// TIA Portal project "oscat_basic_332_s7_TIA_V12_V13_SP1_V14_V15.1" (V15.1)

(* hardware
DEVICE "Rack 0"  S7-300 station
   slot 0: "Profilschiene_0"  Rail  6ES7 390-1***0-0AA0
   slot 2: "Buffer Management"  Unspecific CPU S7 300  6ES7 3XX-XXXXX-XXXX
DEVICE "Rack 0_2"  S7-300 station
   slot 0: "Profilschiene_0"  Rail  6ES7 390-1***0-0AA0
   slot 2: "Constants"  Unspecific CPU S7 300  6ES7 3XX-XXXXX-XXXX
DEVICE "Rack 0_3"  S7-300 station
   slot 0: "Profilschiene_0"  Rail  6ES7 390-1***0-0AA0
   slot 2: "Eng signal generators"  Unspecific CPU S7 300  6ES7 3XX-XXXXX-XXXX
DEVICE "Rack 0_4"  S7-300 station
   slot 0: "Profilschiene_0"  Rail  6ES7 390-1***0-0AA0
   slot 2: "Eng signal processing"  Unspecific CPU S7 300  6ES7 3XX-XXXXX-XXXX
DEVICE "Rack 0_5"  S7-300 station
   slot 0: "Profilschiene_0"  Rail  6ES7 390-1***0-0AA0
   slot 2: "Engineering automation"  Unspecific CPU S7 300  6ES7 3XX-XXXXX-XXXX
DEVICE "Rack 0_6"  S7-300 station
   slot 0: "Profilschiene_0"  Rail  6ES7 390-1***0-0AA0
   slot 2: "Engineering control"  Unspecific CPU S7 300  6ES7 3XX-XXXXX-XXXX
DEVICE "Rack 0_7"  S7-300 station
   slot 0: "Profilschiene_0"  Rail  6ES7 390-1***0-0AA0
   slot 2: "Engineering conversion"  Unspecific CPU S7 300  6ES7 3XX-XXXXX-XXXX
DEVICE "Rack 0_8"  S7-300 station
   slot 0: "Profilschiene_0"  Rail  6ES7 390-1***0-0AA0
   slot 2: "Engineering measurements"  Unspecific CPU S7 300  6ES7 3XX-XXXXX-XXXX
DEVICE "Rack 0_9"  S7-300 station
   slot 0: "Profilschiene_0"  Rail  6ES7 390-1***0-0AA0
   slot 2: "Engineering sensor"  Unspecific CPU S7 300  6ES7 3XX-XXXXX-XXXX
DEVICE "Rack 0_10"  S7-300 station
   slot 0: "Profilschiene_0"  Rail  6ES7 390-1***0-0AA0
   slot 2: "List Processing"  Unspecific CPU S7 300  6ES7 3XX-XXXXX-XXXX
DEVICE "Rack 0_11"  S7-300 station
   slot 0: "Profilschiene_0"  Rail  6ES7 390-1***0-0AA0
   slot 2: "Logic FF edge triggered"  Unspecific CPU S7 300  6ES7 3XX-XXXXX-XXXX
DEVICE "Rack 0_12"  S7-300 station
   slot 0: "Profilschiene_0"  Rail  6ES7 390-1***0-0AA0
   slot 2: "Logic FF pulse triggered"  Unspecific CPU S7 300  6ES7 3XX-XXXXX-XXXX
DEVICE "Rack 0_13"  S7-300 station
   slot 0: "Profilschiene_0"  Rail  6ES7 390-1***0-0AA0
   slot 2: "Logic Others"  Unspecific CPU S7 300  6ES7 3XX-XXXXX-XXXX
DEVICE "Rack 0_14"  S7-300 station
   slot 0: "Profilschiene_0"  Rail  6ES7 390-1***0-0AA0
   slot 2: "Logic gate logic"  Unspecific CPU S7 300  6ES7 3XX-XXXXX-XXXX
DEVICE "Rack 0_15"  S7-300 station
   slot 0: "Profilschiene_0"  Rail  6ES7 390-1***0-0AA0
   slot 2: "Logic generators"  Unspecific CPU S7 300  6ES7 3XX-XXXXX-XXXX
DEVICE "Rack 0_16"  S7-300 station
   slot 0: "Profilschiene_0"  Rail  6ES7 390-1***0-0AA0
   slot 2: "Logic memory"  Unspecific CPU S7 300  6ES7 3XX-XXXXX-XXXX
DEVICE "Rack 0_17"  S7-300 station
   slot 0: "Profilschiene_0"  Rail  6ES7 390-1***0-0AA0
   slot 2: "Math Double Precision"  Unspecific CPU S7 300  6ES7 3XX-XXXXX-XXXX
DEVICE "Rack 0_18"  S7-300 station
   slot 0: "Profilschiene_0"  Rail  6ES7 390-1***0-0AA0
   slot 2: "Math Vektormathematik"  Unspecific CPU S7 300  6ES7 3XX-XXXXX-XXXX
DEVICE "Rack 0_19"  S7-300 station
   slot 0: "Profilschiene_0"  Rail  6ES7 390-1***0-0AA0
   slot 2: "Mathematical"  Unspecific CPU S7 300  6ES7 3XX-XXXXX-XXXX
DEVICE "Rack 0_20"  S7-300 station
   slot 0: "Profilschiene_0"  Rail  6ES7 390-1***0-0AA0
   slot 2: "Mathematical Array"  Unspecific CPU S7 300  6ES7 3XX-XXXXX-XXXX
DEVICE "Rack 0_21"  S7-300 station
   slot 0: "Profilschiene_0"  Rail  6ES7 390-1***0-0AA0
   slot 2: "Mathematical Complex"  Unspecific CPU S7 300  6ES7 3XX-XXXXX-XXXX
DEVICE "Rack 0_22"  S7-300 station
   slot 0: "Profilschiene_0"  Rail  6ES7 390-1***0-0AA0
   slot 2: "Mathematical Geometry"  Unspecific CPU S7 300  6ES7 3XX-XXXXX-XXXX
DEVICE "Rack 0_23"  S7-300 station
   slot 0: "Profilschiene_0"  Rail  6ES7 390-1***0-0AA0
   slot 2: "Mathematical functions"  Unspecific CPU S7 300  6ES7 3XX-XXXXX-XXXX
DEVICE "Rack 0_24"  S7-300 station
   slot 0: "Profilschiene_0"  Rail  6ES7 390-1***0-0AA0
   slot 2: "Other"  Unspecific CPU S7 300  6ES7 3XX-XXXXX-XXXX
DEVICE "Rack 0_25"  S7-300 station
   slot 0: "Profilschiene_0"  Rail  6ES7 390-1***0-0AA0
   slot 2: "String"  Unspecific CPU S7 300  6ES7 3XX-XXXXX-XXXX
DEVICE "Rack 0_26"  S7-300 station
   slot 0: "Profilschiene_0"  Rail  6ES7 390-1***0-0AA0
   slot 2: "Time and Date"  Unspecific CPU S7 300  6ES7 3XX-XXXXX-XXXX
DEVICE "Rack 0_27"  S7-300 station
   slot 0: "Profilschiene_0"  Rail  6ES7 390-1***0-0AA0
   slot 2: "xS7"  Unspecific CPU S7 300  6ES7 3XX-XXXXX-XXXX
*)

// ===== PLC "Buffer Management"  Unspecific CPU S7 300 =====

DATA_BLOCK "SETUP"   // DB1
TITLE = SETUP
{ S7_Optimized_Access := 'FALSE' }
AUTHOR : oscat
FAMILY : CONSTANT
NAME : DBSETUP
VERSION : 1.0
   VAR
      EXTENDED_ASCII : Bool := TRUE;
      CHARNAMES : Array[1..4] of String[253];
      MTH_OFS : Array[1..12] of Int;
      DECADES : Array[0..8] of Real;
   END_VAR
BEGIN
   CHARNAMES[1] := ';"&quot;&&amp;<&lt;>&gt;€&euro; &nbsp;¡&iexcl;¢&cent;£&pound;¤&curren;¥&yen;¦&brvbar;§&sect;¨&uml;©&copy;ª&ordf;«&laquo;¬&not;­&shy;®&reg;¯&macr;°&deg;±&plusmn;²&sup2;³&sup3;´&acute;µ&micro;¶&para;·&middot;¸&cedil;¹&sup1;º&ordm;»&raquo;¼&frac14;Û&Ucirc;';
   CHARNAMES[2] := ';¾&frac34;¿&iquest;À&Agrave;Á&Aacute;Â&Acirc;Ã&Atilde;Ä&Auml;Å&Aring;Æ&AElig;Ç&Ccedil;È&Egrave;É&Eacute;Ê&Ecirc;Ë&Euml;Ì&Igrave;Í&Iacute;Î&Icirc;Ï&Iuml;Ð&ETH;Ñ&Ntilde;Ò&Ograve;Ó&Oacute;Ô&Ocirc;Õ&Otilde;Ö&Ouml;×&times;Ø&Oslash;Ù&Ugrave;Ú&Uacute;½&frac12;';
   CHARNAMES[3] := ';Ü&Uuml;Ý&Yacute;Þ&THORN;ß&szlig;à&agrave;á&aacute;â&acirc;ã&atilde;ä&auml;å&aring;æ&aelig;ç&ccedil;è&egrave;é&eacute;ê&ecirc;ë&euml;ì&igrave;í&iacute;î&icirc;ï&iuml;ð&eth;ñ&ntilde;ò&ograve;ó&oacute;ô&ocirc;õ&otilde;ö&ouml;÷&divide;ø&oslash;ù&ugrave;';
   CHARNAMES[4] := ';ú&uacute;û&ucirc;ü&uuml;ý&yacute;þ&thorn;ÿ&yuml;';
   MTH_OFS[2] := 31;
   MTH_OFS[3] := 59;
   MTH_OFS[4] := 90;
   MTH_OFS[5] := 120;
   MTH_OFS[6] := 151;
   MTH_OFS[7] := 181;
   MTH_OFS[8] := 212;
   MTH_OFS[9] := 243;
   MTH_OFS[10] := 273;
   MTH_OFS[11] := 304;
   MTH_OFS[12] := 334;
   DECADES[0] := 1.0e+0;
   DECADES[1] := 1.0e+1;
   DECADES[2] := 1.0e+2;
   DECADES[3] := 1.0e+3;
   DECADES[4] := 1.0e+4;
   DECADES[5] := 1.0e+4;
   DECADES[6] := 1.0e+5;
   DECADES[7] := 1.0e+6;
   DECADES[8] := 1.0e+7;
END_DATA_BLOCK

FUNCTION_BLOCK "_BUFFER_CLEAR"   // FB225, SCL
TITLE = _BUFFER_CLEAR
{ S7_Optimized_Access := 'FALSE' }
AUTHOR : hugo
FAMILY : BUFFER
NAME : BCLEAR
VERSION : 1.2
// this function will initialize a given array of byte with 0.
// the function needs to be called:    _buffer_clear(adr("array"),sizeof("array"));
// this function will manipulate a given array.
// the function manipulates the original array, it rerturnes true when finished.
// because this function works with pointers its very time efficient and it needs no extra memory.
   VAR_INPUT
      PT : Pointer;
      _PT AT PT : Struct
         DBNr : Word;
         Adr : DWord;
      END_STRUCT;
      SIZE : Int;
   END_VAR
   VAR_OUTPUT
      _CLEAR : Bool;
   END_VAR
   VAR_TEMP
      ptw : Int;   // POINTER TO DWORD;
      temp : DWord;
      end : DWord;
      end32 : DWord;
      tPT : Int;
   END_VAR
BEGIN


   #_CLEAR := FALSE;

   #tPT := DWORD_TO_INT(SHR(IN:=SHL(IN:=#_PT.Adr,N:=8),N:=11));

   (* this routine uses 32 bit access to gain speed *)
   (* first access bytes till pointer is aligned for 32 bit access *)
   #temp := INT_TO_DWORD(#tPT);  //pt;
   #end := DINT_TO_DWORD(DWORD_TO_DINT(#temp) + #SIZE);
   #end32 := DINT_TO_DWORD(DWORD_TO_DINT(#end) - 4);   //end32 := end - 3;
   WHILE (#tPT < DWORD_TO_DINT(#end)) AND (DWORD_TO_DINT((#temp AND 16#00000003)) > 0) DO
       WORD_TO_BLOCK_DB(#_PT.DBNr).DB(#tPT) := 0;
       #tPT := #tPT + 1;
       #temp := DINT_TO_DWORD(DWORD_TO_DINT(#temp) + 1);
   END_WHILE;
   (* pointer is aligned, now copy 32 bits at a time *)
   #ptw := #tPT;
   WHILE #ptw < DWORD_TO_DINT(#end32) DO
       WORD_TO_BLOCK_DB(#_PT.DBNr).DD(#ptw) := 0;
       #ptw := #ptw + 4;
   END_WHILE;
   (* copy the remaining bytes in byte mode *)
   #tPT := #ptw;    //ptw;
   WHILE #tPT < DWORD_TO_DINT(#end) DO
       WORD_TO_BLOCK_DB(#_PT.DBNr).DB(#tPT) := 0;
       #tPT := #tPT + 1;
   END_WHILE;

   #_CLEAR := TRUE;

   (* revision History
   hm  5. mar. 2008    rev 1.0
       original version

   hm  16. mar. 2008   rev 1.1
       added type conversion to avoid warnings under codesys 30
       chaged type of input size to uint
       deleted unused variable i

   hm  31. oct. 2008   rev 1.2
       corrected an error while routine would write outside of arrays

   *)
END_FUNCTION_BLOCK

FUNCTION_BLOCK "_BUFFER_INIT"   // FB226, SCL
TITLE = _BUFFER_INIT
{ S7_Optimized_Access := 'FALSE' }
AUTHOR : hugo
FAMILY : BUFFER
NAME : BINIT
VERSION : 1.2
// this function will initialize a given array of byte with init.
// the function needs to be called:    _buffer_init(adr("array"),sizeof("array"),init);
// this function will manipulate a given array.
// the function manipulates the original array, it rerturnes true when finished.
// because this function works with pointers its very time efficient and it needs no extra memory.
   VAR_INPUT
      pt : Pointer;
      _pt AT pt : Struct
         DBNr : Word;
         Adr : DWord;
      END_STRUCT;
      size : Int;
      init : Byte;
   END_VAR
   VAR_OUTPUT
      _INIT : Bool;
   END_VAR
   VAR_TEMP
      ptw : Int;   // ptw : POINTER TO DWORD;
      temp : DWord;
      end : DWord;
      end32 : DWord;
      tPT : Int;
   END_VAR
BEGIN


   #_INIT := FALSE;
   #tPT := DWORD_TO_INT(SHR(IN:=SHL(IN:=#_pt.Adr,N:=8),N:=11));

   (* this routine uses 32 bit access to gain speed *)
   (* first access bytes till pointer is aligned for 32 bit access *)
   #temp := INT_TO_DWORD(#tPT);
   #end := DINT_TO_DWORD(DWORD_TO_DINT(#temp) + #size);
   #end32 := DINT_TO_DWORD(DWORD_TO_DINT(#temp) - 4);    //end32 := end - 3;
   WHILE (#tPT < DWORD_TO_DINT(#end)) AND (DWORD_TO_DINT((#temp AND 16#00000003)) > 0) DO
       WORD_TO_BLOCK_DB(#_pt.DBNr).DB(#tPT) := #init;
       #tPT := #tPT + 1;
       #temp := DINT_TO_DWORD(DWORD_TO_DINT(#temp) + 1);
   END_WHILE;
   (* pointer is aligned, now copy 32 bits at a time *)
   #ptw := #tPT;
   #temp := SHL(IN:=BYTE_TO_DWORD(#init),N:=24) OR SHL(IN:=BYTE_TO_DWORD(#init),N:=16) OR SHL(IN:=BYTE_TO_DWORD(#init),N:=8) OR BYTE_TO_DWORD(#init);
   WHILE #ptw < DWORD_TO_DINT(#end32) DO
       WORD_TO_BLOCK_DB(#_pt.DBNr).DD(#ptw) := #temp;
       #ptw := #ptw + 4;
   END_WHILE;
   (* copy the remaining bytes in byte mode *)
   #tPT := #ptw;
   WHILE #tPT < DWORD_TO_DINT(#end) DO
       WORD_TO_BLOCK_DB(#_pt.DBNr).DB(#tPT) := #init;
       #tPT := #tPT + 1;
   END_WHILE;

   #_INIT := TRUE;

   (* revision History
   hm  5. mar. 2008    rev 1.0
       original version

   hm  16. mar. 2008   rev 1.1
       added type conversion to avoid warnings under codesys 3.0
       chaged type of input size to uint.

   hm  31. oct. 2008   rev 1.2
       corrected an error while routine would write outside of arrays

   *)
END_FUNCTION_BLOCK

FUNCTION_BLOCK "_BUFFER_INSERT"   // FB227, SCL
TITLE = _BUFFER_INSERT
{ S7_Optimized_Access := 'FALSE' }
AUTHOR : hugo
FAMILY : BUFFER
NAME : BINSERT
VERSION : 1.4
// this function will initialize a given array of byte with init.
// the function needs to be called:    _buffer_init(adr("array"),sizeof("array"),init);
// this function will manipulate a given array.
// the function manipulates the original array, it rerturnes true when finished.
// because this function works with pointers its very time efficient and it needs no extra memory.
// 
// uses: STRING_TO_BUFFER [FB228]
   VAR_INPUT
      STR : String[254];
      _str AT STR : Struct
         length : Byte;
         act_length : Byte;
         str : Array[1..254] of Byte;
      END_STRUCT;
      POS : Int;
      PT : Pointer;
      _pt AT PT : Struct
         DBNr : Word;
         Adr : DWord;
      END_STRUCT;
      SIZE : Int;
   END_VAR
   VAR_OUTPUT
      OUT : Bool;
   END_VAR
   VAR
      STRING_TO_BUFFER : "_STRING_TO_BUFFER";
   END_VAR
   VAR_TEMP
      end : Int;
      lx : Int;
      i : Int;
      tPT : Int;
   END_VAR
BEGIN


   #OUT := FALSE;

   #tPT := DWORD_TO_INT(SHR(IN:=SHL(IN:=#_pt.Adr,N:=8),N:=11));

   #POS := LIMIT(MN:=0,IN:=#POS,MX:=#SIZE - 1);
   #lx := BYTE_TO_INT(#_str.length);  //LEN(str);
   #end := #POS + #lx;
   (* first move the upper part of the buffer to make space for the string *)
   FOR #i := #SIZE - 1 TO #end BY -1 DO
       WORD_TO_BLOCK_DB(#_pt.DBNr).DB(#tPT+#i) := WORD_TO_BLOCK_DB(#_pt.DBNr).DB(#tPT+#i-#lx);
   END_FOR;
   (* copy the string *)
   #STRING_TO_BUFFER(strBLKMOV#STR, pos:=#POS, pt:=#PT, size:=#SIZE);
   #OUT := #STRING_TO_BUFFER._BUFFER;


   (* revision History
   hm  9. mar. 2008  rev 1.0
     original version

   hm  16. mar. 2008 rev 1.1
     changed type of input size to uint

   hm  13. may. 2008 rev 1.2
     changed type of pointer to array[1..32767]
     changed size of string to STRING_LENGTH

   hm  23. mar. 2009 rev 1.3
     avoid writing to input pos

   hm  12. nov. 2009 rev 1.4
     code optimized

   *)
END_FUNCTION_BLOCK

FUNCTION_BLOCK "_STRING_TO_BUFFER"   // FB228, SCL
TITLE = _STRING_TO_BUFFER
{ S7_Optimized_Access := 'FALSE' }
AUTHOR : hugo
FAMILY : BUFFER
NAME : BSTRB
VERSION : 1.3
// this function will copy a string into an array of byte starting at position pos.
// the function needs to be called:    _String_To_buffer(str, pos, adr("array"),sizeof("array"));
// this function will manipulate the array directly in memory and returns true when finished.
// because this function works with pointers its very time efficient and it needs no extra memory.
   VAR_INPUT
      str : String[254];
      _str AT str : Struct
         length : Byte;
         act_length : Byte;
         str : Array[1..254] of Byte;
      END_STRUCT;
      pos : Int;
      pt : Pointer;
      _pt AT pt : Struct
         DBNr : Word;
         Adr : DWord;
      END_STRUCT;
      size : Int;
   END_VAR
   VAR_OUTPUT
      _BUFFER : Bool;
   END_VAR
   VAR_TEMP
      ps : Int;   // POINTER TO BYTE;
      i : Int;
      end : Int;
      tPT : Int;
   END_VAR
BEGIN


   #_BUFFER := FALSE;
   #tPT := DWORD_TO_INT(SHR(IN:=SHL(IN:=#_pt.Adr,N:=8),N:=11));

   #ps := 1;    //ADR(str);
   #end := MIN(IN1:=#pos + BYTE_TO_INT(#_str.length) - 1,IN2:=#size);
   IF #end > 0 THEN #end := #end -1; END_IF;
   FOR #i := #pos TO #end DO
       WORD_TO_BLOCK_DB(#_pt.DBNr).DB(#tPT+#i-1) := #_str.str[#ps];
       #ps := #ps + 1;
   END_FOR;

   #_BUFFER := TRUE;

   (* revision History

   hm  5. mar. 2008 rev 1.0
    original version

   hm 16. mar. 2008 rev 1.1
    changed type of input size to uint

   hm 13. may. 2008 rev 1.2
    changed type of pointer to array[1..32767]
    changed size of string to STRING_LENGTH

   hm 12. nov. 2009 rev 1.3
    limit end to size - 1

   *)
END_FUNCTION_BLOCK

FUNCTION_BLOCK "BUFFER_SEARCH"   // FB229, SCL
TITLE = BUFFER_SEARCH
{ S7_Optimized_Access := 'FALSE' }
AUTHOR : hugo
FAMILY : BUFFER
NAME : BSEARCH
VERSION : 1.4
// this function will search for a string STR in an array of byte starting at position pos.
// the function needs to be called: buffer_search(adr("array"),sizeof("array"), STR, POS, IGN);
// because this function works with pointers its very time efficient and it needs no extra memory.
// The function returns the position of the first character of the string in the array if found.
// a -1 is returned if the string is not found in the array.
// when IGN = TRUE, STR must be in capital letters and the search is case insensitv.
   VAR_INPUT
      PT : Pointer;
      _pt AT PT : Struct
         DBNr : Word;
         Adr : DWord;
      END_STRUCT;
      SIZE : Int;
      STR : String[254];
      _str AT STR : Struct
         length : Byte;
         act_length : Byte;
         str : Array[1..254] of Byte;
      END_STRUCT;
      POS : Int;
      IGN : Bool;
   END_VAR
   VAR_OUTPUT
      _SEARCH : Int;
   END_VAR
   VAR_TEMP
      ps : Int;   // POINTER TO ARRAY[0..255] OF BYTE;
      chx : Byte;
      i : Int;
      end : Int;
      k : Int;
      lx : Int;
      tPT : Int;
   END_VAR
BEGIN


   #tPT := DWORD_TO_INT(SHR(IN:=SHL(IN:=#_pt.Adr,N:=8),N:=11));

   #ps := 1;    //ADR(str);
   #lx := BYTE_TO_INT(#_str.act_length);  //LEN(str);
   #end := MIN(IN1:=#SIZE - #lx, IN2:= #SIZE - 1);
   #lx := #lx - 1;
   FOR #i := #POS TO #end DO
     FOR #k := 0 TO #lx DO
       //IF (_str.str[ps+k] <> ign) AND (_str.str[ps+k] <> WORD_TO_BLOCK_DB(_pt.DBNr).DB[tPT+i+k]) THEN EXIT; END_IF;
       IF #IGN THEN 
         #chx := "TO_UPPER"(WORD_TO_BLOCK_DB(#_pt.DBNr).DB(#tPT+#i+#k)); 
       ELSE 
         #chx := WORD_TO_BLOCK_DB(#_pt.DBNr).DB(#tPT+#i+#k); 
       END_IF;
       IF WORD_TO_BLOCK_DB(#_pt.DBNr).DB(#tPT+#k) <> #chx THEN 
         EXIT; 
       END_IF;
     END_FOR;
     IF #k > #lx THEN
       #_SEARCH := #i;
       RETURN;
     END_IF;
   END_FOR;
   #_SEARCH := -1;


   (* revision History

   hm 5. mar. 2008 rev 1.0
     original version

   hm  16. mar. 2008 rev 1.1
     chaged type of input size to uint

   hm  13. may. 2008 rev 1.2
     changed type of pointer to array[1..32767]
     changed size of string to STRING_LENGTH

   hm  12. nov. 2009 rev 1.3
     limit end to array size

   hm  25. jan. 2011 rev 1.4
     ign = True will now ignore case
     return -1 if nothing found
   *)
END_FUNCTION_BLOCK

FUNCTION_BLOCK "BUFFER_TO_STRING"   // FB230, SCL
TITLE = BUFFER_TO_STRING
{ S7_Optimized_Access := 'FALSE' }
AUTHOR : hugo
FAMILY : BUFFER
NAME : BBSTR
VERSION : 1.5
// this function will retrieve a string from an array of byte starting at position start and stop at position stop.
// the function needs to be called: buffer_TO_String(adr("array"),sizeof("array"), start, stop);
// because this function works with pointers its very time efficient and it needs no extra memory.
   VAR_INPUT
      PT : Pointer;
      _pt AT PT : Struct
         DBNr : Word;
         Adr : DWord;
      END_STRUCT;
      SIZE : Int;
      START : Int;
      STOP : Int;
   END_VAR
   VAR_OUTPUT
      _STRING : String[254];
      _str AT _STRING : Struct
         length : Byte;
         act_length : Byte;
         str : Array[1..254] of Byte;
      END_STRUCT;
   END_VAR
   VAR_TEMP
      ps : Int;   // POINTER TO BYTE;
      i : Int;
      tPT : Int;
      stp : Int;
      sta : Int;
   END_VAR
BEGIN


   #tPT := DWORD_TO_INT(SHR(IN:=SHL(IN:=#_pt.Adr,N:=8),N:=11));

   #ps := 1;    //ADR(BUFFER_TO_STRING);
   IF #SIZE = 0 THEN RETURN; END_IF;
   #sta := MIN(IN1:=#START, IN2:=#SIZE-1);
   #stp := MIN(IN1:=#STOP, IN2:=#SIZE-1);

   (* check for maximum string_length *)
   IF (#stp - #sta + 1) >= BYTE_TO_INT(#_str.act_length) THEN
     #stp := #sta + BYTE_TO_INT(#_str.act_length) - 1;
   END_IF;

   FOR #i := #sta TO #stp DO
       #_str.str[#ps] := WORD_TO_BLOCK_DB(#_pt.DBNr).DB(#tPT+#i);
       #ps := #ps + 1;
   END_FOR;

   (* terminate the string *)
   #_str.act_length := INT_TO_BYTE(#ps-1);

   (* revision History
   hm  5. mar. 2008  rev 1.0
     original version

   hm  16. mar. 2008 rev 1.1
     changed type of input size to uint

   hm  13. may. 2008 rev 1.2
     changed type of pointer to array[0..32767]
     changed size of string to STRING_LENGTH

   hm  12. jun. 2008 rev 1.3
     check for pointer overrun
     change input start and stop to uint
     added type conversions to avoid warnings under codesys 3.0

   hm  23. mar. 2009 rev 1.4
     avoid writing to input stop

   hm  12. nov. 2009 rev 1.5
     limit start and stop to size -1

   *)
END_FUNCTION_BLOCK

FUNCTION_BLOCK "BUFFER_COMP"   // FB243, SCL
TITLE = BUFFER_COMP
{ S7_Optimized_Access := 'FALSE' }
AUTHOR : hugo
FAMILY : BUFFER
NAME : BCOMP
VERSION : 1.1
   VAR_INPUT
      PT1 : Pointer;   // POINTER TO ARRAY OF BYTE
      _PT1 AT PT1 : Struct
         DBNr : Word;
         Adr : DWord;
      END_STRUCT;
      SIZE1 : Int;
      PT2 : Pointer;   // POINTER TO ARRAY OF BYTE
      _PT2 AT PT2 : Struct
         DBNr : Word;
         Adr : DWord;
      END_STRUCT;
      SIZE2 : Int;
      START : Int;
   END_VAR
   VAR_OUTPUT
      COMP : Int;
   END_VAR
   VAR
      i : Int;
      j : Int;
      end : Int;
      firstbyte : Byte;
   END_VAR
   VAR_TEMP
      tPT1 : Int;
      tPT2 : Int;
   END_VAR
BEGIN

   //WORD_TO_BLOCK_DB(_pt.DBNr).DB[tPT+i+k-1])
   #COMP := 0;

   (* get start address of pointer *)
   #tPT1 := DWORD_TO_INT(SHR(IN:=SHL(IN:=#_PT1.Adr,N:=8),N:=11));
   #tPT2 := DWORD_TO_INT(SHR(IN:=SHL(IN:=#_PT2.Adr,N:=8),N:=11));

   (* search for first character match *)
   IF #SIZE2 <= #SIZE1 THEN
       #end := #SIZE1 - #SIZE2;
       #firstbyte := WORD_TO_BLOCK_DB(#_PT2.DBNr).DB(#tPT2);
       FOR #i := #START TO #end DO
           IF WORD_TO_BLOCK_DB(#_PT1.DBNr).DB(#tPT1+#i) = #firstbyte THEN
               (* first character matches, now compare rest of array *)
               #j := 1;
               WHILE #j < #SIZE2 DO
                   IF WORD_TO_BLOCK_DB(#_PT2.DBNr).DB(#tPT2+#j) <> WORD_TO_BLOCK_DB(#_PT1.DBNr).DB(#tPT1+#j+#i) THEN EXIT; END_IF;
                   #j := #j + 1;
               END_WHILE;
               (* when J > size2 a match was found return the position i in buffer1 *)
               IF #j = #SIZE2 THEN
                   #COMP := #i;
                   RETURN;
               END_IF;
           END_IF;
       END_FOR;
   END_IF;
   #COMP := -1;


   (*
   hm 14. nov. 2008  rev 1.0
     original version

   hm  12. nov. 2009 rev 1.1
     performance increase

   *)
END_FUNCTION_BLOCK

FUNCTION_BLOCK "_BUFFER_UPPERCASE"   // FB255, SCL
TITLE = _BUFFER_UPPERCASE
{ S7_Optimized_Access := 'FALSE' }
AUTHOR : hugo
FAMILY : BUFFER
NAME : BUPPER
VERSION : 1.0
// this FUNCTION will convert an ARRAY OF BYTE into uppercase
// the function needs to be called:  _buffer_clear(adr("array"),sizeof("array"));
// this function will manipulate a given array.
// the function manipulates the original array, it rerturnes true when finished.
// because this function works with pointers its very time efficient and it needs no extra memory.
   VAR_INPUT
      PT : Pointer;
      _PT AT PT : Struct
         DBNr : Word;
         Adr : DWord;
      END_STRUCT;
      SIZE : Int;
   END_VAR
   VAR_OUTPUT
      UPPERCASE : Bool;
   END_VAR
   VAR_TEMP
      pos : Int;
      tPT : Int;
   END_VAR
BEGIN


   #UPPERCASE := FALSE;

   #tPT := DWORD_TO_INT(SHR(IN:=SHL(IN:=#_PT.Adr,N:=8),N:=11));

   #pos := 0;
   WHILE #pos < #SIZE DO
     WORD_TO_BLOCK_DB(#_PT.DBNr).DB(#tPT+#pos) := "TO_UPPER"(WORD_TO_BLOCK_DB(#_PT.DBNr).DB(#tPT+#pos));
     #pos := #pos + 1;
   END_WHILE;

   #UPPERCASE := TRUE;


   (* revision History
   hm  20. jan. 2011 rev 1.0
     original version

   *)
END_FUNCTION_BLOCK

FUNCTION "TO_UPPER" : Byte   // FC284, SCL
TITLE = TO_UPPER
{ S7_Optimized_Access := 'FALSE' }
AUTHOR : hugo
FAMILY : STRINGS
NAME : TO_UPPER
VERSION : 1.3
// to_upper converts a character from lowercase to uppercase
// 
// uses: SETUP [DB1]
   VAR_INPUT
      IN : Byte;
   END_VAR
BEGIN


   IF BYTE_TO_INT(#IN) > 96 AND BYTE_TO_INT(#IN) < 123 THEN
      #TO_UPPER := #IN AND 16#DF;
   ELSIF BYTE_TO_INT(#IN) > 223 AND BYTE_TO_INT(#IN) <> 247 AND BYTE_TO_INT(#IN) <> 255 AND "SETUP".EXTENDED_ASCII THEN
      #TO_UPPER := #IN AND 16#DF;
   ELSE
      #TO_UPPER := #IN;
   END_IF;


   (* revision history
   hm  6. mar. 2008    rev 1.0
       original version

   hm  19. oct. 2008   rev 1.1
       changed setup constants

   ks  25. oct. 2008   rev 1.2
       optimized code

   hm 16. jan 2009 rev 1.3
       corrected an error in module

   *)
END_FUNCTION

// ===== PLC "Constants"  Unspecific CPU S7 300 =====

DATA_BLOCK "SETUP"   // DB1
TITLE = SETUP
{ S7_Optimized_Access := 'FALSE' }
AUTHOR : oscat
FAMILY : CONSTANT
NAME : DBSETUP
VERSION : 1.0
   VAR
      EXTENDED_ASCII : Bool := TRUE;
      CHARNAMES : Array[1..4] of String[253];
      MTH_OFS : Array[1..12] of Int;
      DECADES : Array[0..8] of Real;
   END_VAR
BEGIN
   CHARNAMES[1] := ';"&quot;&&amp;<&lt;>&gt;€&euro; &nbsp;¡&iexcl;¢&cent;£&pound;¤&curren;¥&yen;¦&brvbar;§&sect;¨&uml;©&copy;ª&ordf;«&laquo;¬&not;­&shy;®&reg;¯&macr;°&deg;±&plusmn;²&sup2;³&sup3;´&acute;µ&micro;¶&para;·&middot;¸&cedil;¹&sup1;º&ordm;»&raquo;¼&frac14;Û&Ucirc;';
   CHARNAMES[2] := ';¾&frac34;¿&iquest;À&Agrave;Á&Aacute;Â&Acirc;Ã&Atilde;Ä&Auml;Å&Aring;Æ&AElig;Ç&Ccedil;È&Egrave;É&Eacute;Ê&Ecirc;Ë&Euml;Ì&Igrave;Í&Iacute;Î&Icirc;Ï&Iuml;Ð&ETH;Ñ&Ntilde;Ò&Ograve;Ó&Oacute;Ô&Ocirc;Õ&Otilde;Ö&Ouml;×&times;Ø&Oslash;Ù&Ugrave;Ú&Uacute;½&frac12;';
   CHARNAMES[3] := ';Ü&Uuml;Ý&Yacute;Þ&THORN;ß&szlig;à&agrave;á&aacute;â&acirc;ã&atilde;ä&auml;å&aring;æ&aelig;ç&ccedil;è&egrave;é&eacute;ê&ecirc;ë&euml;ì&igrave;í&iacute;î&icirc;ï&iuml;ð&eth;ñ&ntilde;ò&ograve;ó&oacute;ô&ocirc;õ&otilde;ö&ouml;÷&divide;ø&oslash;ù&ugrave;';
   CHARNAMES[4] := ';ú&uacute;û&ucirc;ü&uuml;ý&yacute;þ&thorn;ÿ&yuml;';
   MTH_OFS[2] := 31;
   MTH_OFS[3] := 59;
   MTH_OFS[4] := 90;
   MTH_OFS[5] := 120;
   MTH_OFS[6] := 151;
   MTH_OFS[7] := 181;
   MTH_OFS[8] := 212;
   MTH_OFS[9] := 243;
   MTH_OFS[10] := 273;
   MTH_OFS[11] := 304;
   MTH_OFS[12] := 334;
   DECADES[0] := 1.0e+0;
   DECADES[1] := 1.0e+1;
   DECADES[2] := 1.0e+2;
   DECADES[3] := 1.0e+3;
   DECADES[4] := 1.0e+4;
   DECADES[5] := 1.0e+4;
   DECADES[6] := 1.0e+5;
   DECADES[7] := 1.0e+6;
   DECADES[8] := 1.0e+7;
END_DATA_BLOCK

DATA_BLOCK "MATH"   // DB2
TITLE = MATH
{ S7_Optimized_Access := 'FALSE' }
AUTHOR : oscat
FAMILY : CONSTANT
NAME : DBMATH
VERSION : 1.1
   VAR
      PI : Real := 3.141593e+0;   // Kreiszahl PI
      PI2 : Real := 6.283185e+0;   // PI * 2
      PI4 : Real := 1.256637e+1;   // PI * 4
      PI05 : Real := 1.570796e+0;   // PI / 2
      PI025 : Real := 7.853982e-1;   // PI / 4
      PI_INV : Real := 3.183099e-1;   // 1 / PI
      "E" : Real := 2.718282e+0;   // Eulersche Konstante
      E_INV : Real := 3.678795e-1;   // 1 / e
      SQ2 : Real := 1.414214e+0;   // Wurzel von 2
      FACTS : Array[0..12] of DInt;
   END_VAR
BEGIN
   FACTS[0] := DINT#1;
   FACTS[1] := DINT#1;
   FACTS[2] := DINT#2;
   FACTS[3] := DINT#6;
   FACTS[4] := DINT#24;
   FACTS[5] := DINT#120;
   FACTS[6] := DINT#720;
   FACTS[7] := DINT#5040;
   FACTS[8] := DINT#40320;
   FACTS[9] := DINT#362880;
   FACTS[10] := DINT#3628800;
   FACTS[11] := DINT#39916800;
   FACTS[12] := DINT#479001600;
END_DATA_BLOCK

DATA_BLOCK "PHYS"   // DB3
TITLE = PHYS
{ S7_Optimized_Access := 'FALSE' }
AUTHOR : oscat
FAMILY : CONSTANT
NAME : DBPHYS
VERSION : 1.1
// CONSTANTS_PHYS
   VAR
      C : Real := 2.997924e+8;   // Lichtgeschwindigkeit in m/s
      "E" : Real := 1.602176e-19;   // elementarladung in Colomb = A * s
      G : Real := 9.80665e+0;   // Erdbeschleunigung in m / s²
      T0 : Real := -2.7315e+2;   // absoluter Nullpunkt in °C
      RU : Real := 8.314472e+0;   // Universelle Gaskonstante in J / (mol · K)
      PN : Real := 1.01325e+5;   // NormalDruck in Pa
   END_VAR
BEGIN
END_DATA_BLOCK

DATA_BLOCK "LANGUAGE"   // DB4
TITLE = LANGUAGE
{ S7_Optimized_Access := 'FALSE' }
AUTHOR : oscat
FAMILY : CONSTANT
NAME : DBLANG
VERSION : 1.2
   VAR
      DEFAULT : Int := 1;   // 1=english, 2=german, 3=french
      LMAX : Int := 3;
      WEEKDAYS : Array[1..3, 1..7] of String[10];
      WEEKDAYS2 : Array[1..3, 1..7] of String[2];
      MONTHS : Array[1..3, 1..12] of String[10];
      MONTHS3 : Array[1..3, 1..12] of String[3];
      DIRS : Array[1..3, 0..15] of String[3];
   END_VAR
BEGIN
   WEEKDAYS[1,1] := 'Monday';
   WEEKDAYS[1,2] := 'Tuesday';
   WEEKDAYS[1,3] := 'Wednesday';
   WEEKDAYS[1,4] := 'Thursday';
   WEEKDAYS[1,5] := 'Friday';
   WEEKDAYS[1,6] := 'Saturday';
   WEEKDAYS[1,7] := 'Sunday';
   WEEKDAYS[2,1] := 'Montag';
   WEEKDAYS[2,2] := 'Dienstag';
   WEEKDAYS[2,3] := 'Mittwoch';
   WEEKDAYS[2,4] := 'Donnerstag';
   WEEKDAYS[2,5] := 'Freitag';
   WEEKDAYS[2,6] := 'Samstag';
   WEEKDAYS[2,7] := 'Sonntag';
   WEEKDAYS[3,1] := 'Lundi';
   WEEKDAYS[3,2] := 'Mardi';
   WEEKDAYS[3,3] := 'Mercredi';
   WEEKDAYS[3,4] := 'Jeudi';
   WEEKDAYS[3,5] := 'Vendredi';
   WEEKDAYS[3,6] := 'Samedi';
   WEEKDAYS[3,7] := 'Dimanche';
   WEEKDAYS2[1,1] := 'Mo';
   WEEKDAYS2[1,2] := 'Tu';
   WEEKDAYS2[1,3] := 'We';
   WEEKDAYS2[1,4] := 'Th';
   WEEKDAYS2[1,5] := 'Fr';
   WEEKDAYS2[1,6] := 'Sa';
   WEEKDAYS2[1,7] := 'Su';
   WEEKDAYS2[2,1] := 'Mo';
   WEEKDAYS2[2,2] := 'Di';
   WEEKDAYS2[2,3] := 'Mi';
   WEEKDAYS2[2,4] := 'Do';
   WEEKDAYS2[2,5] := 'Fr';
   WEEKDAYS2[2,6] := 'Sa';
   WEEKDAYS2[2,7] := 'So';
   WEEKDAYS2[3,1] := 'Lu';
   WEEKDAYS2[3,2] := 'Ma';
   WEEKDAYS2[3,3] := 'Me';
   WEEKDAYS2[3,4] := 'Je';
   WEEKDAYS2[3,5] := 'Ve';
   WEEKDAYS2[3,6] := 'Sa';
   WEEKDAYS2[3,7] := 'Di';
   MONTHS[1,1] := 'January';
   MONTHS[1,2] := 'February';
   MONTHS[1,3] := 'March';
   MONTHS[1,4] := 'April';
   MONTHS[1,5] := 'May';
   MONTHS[1,6] := 'June';
   MONTHS[1,7] := 'July';
   MONTHS[1,8] := 'August';
   MONTHS[1,9] := 'September';
   MONTHS[1,10] := 'October';
   MONTHS[1,11] := 'November';
   MONTHS[1,12] := 'December';
   MONTHS[2,1] := 'Januar';
   MONTHS[2,2] := 'Februar';
   MONTHS[2,3] := 'März';
   MONTHS[2,4] := 'April';
   MONTHS[2,5] := 'Mai';
   MONTHS[2,6] := 'Juni';
   MONTHS[2,7] := 'Juli';
   MONTHS[2,8] := 'August';
   MONTHS[2,9] := 'September';
   MONTHS[2,10] := 'Oktober';
   MONTHS[2,11] := 'November';
   MONTHS[2,12] := 'Dezember';
   MONTHS[3,1] := 'Janvier';
   MONTHS[3,2] := 'Février';
   MONTHS[3,3] := 'mars';
   MONTHS[3,4] := 'Avril';
   MONTHS[3,5] := 'Mai';
   MONTHS[3,6] := 'Juin';
   MONTHS[3,7] := 'Juillet';
   MONTHS[3,8] := 'Août';
   MONTHS[3,9] := 'Septembre';
   MONTHS[3,10] := 'Octobre';
   MONTHS[3,11] := 'Novembre';
   MONTHS[3,12] := 'Decembre';
   MONTHS3[1,1] := 'Jan';
   MONTHS3[1,2] := 'Feb';
   MONTHS3[1,3] := 'Mar';
   MONTHS3[1,4] := 'Apr';
   MONTHS3[1,5] := 'May';
   MONTHS3[1,6] := 'Jun';
   MONTHS3[1,7] := 'Jul';
   MONTHS3[1,8] := 'Aug';
   MONTHS3[1,9] := 'Sep';
   MONTHS3[1,10] := 'Oct';
   MONTHS3[1,11] := 'Nov';
   MONTHS3[1,12] := 'Dec';
   MONTHS3[2,1] := 'Jan';
   MONTHS3[2,2] := 'Feb';
   MONTHS3[2,3] := 'Mrz';
   MONTHS3[2,4] := 'Apr';
   MONTHS3[2,5] := 'Mai';
   MONTHS3[2,6] := 'Jun';
   MONTHS3[2,7] := 'Jul';
   MONTHS3[2,8] := 'Aug';
   MONTHS3[2,9] := 'Sep';
   MONTHS3[2,10] := 'Okt';
   MONTHS3[2,11] := 'Nov';
   MONTHS3[2,12] := 'Dez';
   MONTHS3[3,1] := 'Jan';
   MONTHS3[3,2] := 'Fev';
   MONTHS3[3,3] := 'Mar';
   MONTHS3[3,4] := 'Avr';
   MONTHS3[3,5] := 'Mai';
   MONTHS3[3,6] := 'Jun';
   MONTHS3[3,7] := 'Jul';
   MONTHS3[3,8] := 'Aou';
   MONTHS3[3,9] := 'Sep';
   MONTHS3[3,10] := 'Oct';
   MONTHS3[3,11] := 'Nov';
   MONTHS3[3,12] := 'Dec';
   DIRS[1,0] := 'N';
   DIRS[1,1] := 'NNE';
   DIRS[1,2] := 'NE';
   DIRS[1,3] := 'ENE';
   DIRS[1,4] := 'E';
   DIRS[1,5] := 'ESE';
   DIRS[1,6] := 'SE';
   DIRS[1,7] := 'SSE';
   DIRS[1,8] := 'S';
   DIRS[1,9] := 'SSW';
   DIRS[1,10] := 'SW';
   DIRS[1,11] := 'WSW';
   DIRS[1,12] := 'W';
   DIRS[1,13] := 'WNW';
   DIRS[1,14] := 'NW';
   DIRS[1,15] := 'NNW';
   DIRS[2,0] := 'N';
   DIRS[2,1] := 'NNO';
   DIRS[2,2] := 'NO';
   DIRS[2,3] := 'ONO';
   DIRS[2,4] := 'O';
   DIRS[2,5] := 'OSO';
   DIRS[2,6] := 'SO';
   DIRS[2,7] := 'SSO';
   DIRS[2,8] := 'S';
   DIRS[2,9] := 'SSW';
   DIRS[2,10] := 'SW';
   DIRS[2,11] := 'WSW';
   DIRS[2,12] := 'W';
   DIRS[2,13] := 'WNW';
   DIRS[2,14] := 'NW';
   DIRS[2,15] := 'NNW';
   DIRS[3,0] := 'N';
   DIRS[3,1] := 'NNO';
   DIRS[3,2] := 'NO';
   DIRS[3,3] := 'ONO';
   DIRS[3,4] := 'O';
   DIRS[3,5] := 'OSO';
   DIRS[3,6] := 'SO';
   DIRS[3,7] := 'SSO';
   DIRS[3,8] := 'S';
   DIRS[3,9] := 'SSW';
   DIRS[3,10] := 'SW';
   DIRS[3,11] := 'WSW';
   DIRS[3,12] := 'W';
   DIRS[3,13] := 'WNW';
   DIRS[3,14] := 'NW';
   DIRS[3,15] := 'NNW';
END_DATA_BLOCK

DATA_BLOCK "LOCATION"   // DB5
TITLE = LOCATION
{ S7_Optimized_Access := 'FALSE' }
AUTHOR : oscat
FAMILY : CONSTANT
NAME : DBLOCA
VERSION : 1.2
   VAR
      DEFAULT : Int := 1;   // 1=germany, 2=austria 3=france 4=belgium-german 5= italien-Südtirol
      LMAX : Int := 5;   // language spoken in the location
      LANGUAGE : Array[1..5] of Int;
   END_VAR
BEGIN
   LANGUAGE[1] := 2;
   LANGUAGE[2] := 2;
   LANGUAGE[3] := 3;
   LANGUAGE[4] := 2;
   LANGUAGE[5] := 2;
END_DATA_BLOCK

DATA_BLOCK "CONSTANTS"   // DB6
TITLE = CONSTANTS
{ S7_Optimized_Access := 'FALSE' }
AUTHOR : oscat
FAMILY : CONSTANT
NAME : CONSTANT
VERSION : 1.0
   VAR
      STRING_LENGTH : Int := 250;
      LIST_LENGTH : Int := 250;
   END_VAR
BEGIN
END_DATA_BLOCK

// ===== PLC "Eng signal generators"  Unspecific CPU S7 300 =====

VAR_GLOBAL CONSTANT   // PLC tag table "STEP7 classic symbols"
   "debug" : Bool := FALSE;
   "N" : Int := 0;
   "offset" : Int := 0;
   "E" : Real := 2.71828182845904523536028747135266249;   // Eulersche Konstante
   "PI2" : Real := 6.28318530717958647692528676655900576;   // PI * 2
   "offset_1" : DWord := 0;
END_VAR

DATA_BLOCK "IDB_STIME"   // DB64
{ S7_Optimized_Access := 'FALSE' }
AUTHOR : dalbi
FAMILY : MEASURE
VERSION : 0.0
// stored: InstanceOfName STIME
"STIME"
BEGIN
END_DATA_BLOCK

FUNCTION_BLOCK "CLK_PRG"   // FB52, SCL
TITLE = CLK_PRG
{ S7_Optimized_Access := 'FALSE' }
AUTHOR : hugo
FAMILY : GENERAT
NAME : CLK_PRG
VERSION : 1.3
// clk_prg uses the internal sps time to generate a clock with programmable period time.
// the period time is defined for 10ms .. 65s
// the first cycle after start is a clk pulse and then depending on the programmed period time a delay.
// every pulse is only valid for one cycle.
// the accuracy of clk_prg is depending on the accuracy of the system clock.
// 
// uses: T_PLC_MS [FC64]
//       STIME [FB64],IDB_STIME [DB64]
   VAR_INPUT
      PT : Time := T#10MS;
   END_VAR
   VAR_OUTPUT
      Q : Bool;
   END_VAR
   VAR
      init : Bool;
      last : Time;
      tx : Time;
   END_VAR
   VAR_TEMP
      TOP_SI : Struct
         EV_CLASS : Byte;
         EV_NUM : Byte;
         PRIORITY : Byte;
         NUM : Byte;
         TYP2_3 : Byte;
         TYP1 : Byte;
         ZI1 : Word;
         ZI2_3 : DWord;
      END_STRUCT;
      START_UP_SI : Struct
         EV_CLASS : Byte;
         EV_NUM : Byte;
         PRIORITY : Byte;
         NUM : Byte;
         TYP2_3 : Byte;
         TYP1 : Byte;
         ZI1 : Word;
         ZI2_3 : DWord;
      END_STRUCT;
      ERR : Int;
   END_VAR
BEGIN


   (* read actual startup info *)
   (* OB1_SCAN_1  BYTE  -  B#16#01: Abschluss des Neustarts (Warmstarts)
                        -  B#16#02: Abschluss des Wiederanlaufs
                        -  B#16#03: Abschluss des freien Zyklus
                        -  B#16#04: Abschluss des Kaltstarts
                        -  B#16#05: Erster OB 1-Zyklus der neuen Master-CPU nach 
                                    Master-Reserve-Umschaltung und STOP des 
                                    bisherigen Masters *)

   #ERR := RD_SINFO (TOP_SI => #TOP_SI, START_UP_SI => #START_UP_SI);

   (* read system time *)
   #tx := T_CONV(DWORD_TO_DINT("T_PLC_MS"()));

   (* reset last_time on system startup *)
   IF #TOP_SI.EV_NUM = 1 OR #TOP_SI.EV_NUM = 2 OR #TOP_SI.EV_NUM = 4 THEN 
       #init := false;
   END_IF;

   (* initialize on startup *)
   IF NOT #init THEN
       #init := TRUE;
       #last := #tx - #PT;
   END_IF;

   (* generate output pulse when next_pulse is reached *)
   #Q := #tx - #last >= #PT;
   IF #Q THEN #last := #tx; END_IF;


   (* revision hiostory

   hm 25 feb 2007  rev 1.1
       rewritten code for higher performance
       pt can now be changed during runtime

   hm  17. sep 2007    rev 1.2
       replaced time() with t_plc_ms() for compatibility reasons

   hm  25. oct. 2008   rev 1.3
       optimized code

   *)
END_FUNCTION_BLOCK

FUNCTION_BLOCK "STIME"   // FB64, SCL
TITLE = STIME
{ S7_Optimized_Access := 'FALSE' }
AUTHOR : dalbi
FAMILY : MEASURE
NAME : STIME
VERSION : 1.5
// this function block makes sure that the timer of a siemens sps counts from 0 - 2^32-1.
   VAR_OUTPUT
      tx : DWord;
      at_tx AT tx : Array[0..31] of Bool;
   END_VAR
   VAR
      last_time : DWord;
      bit31 : Bool;
      init : Bool := TRUE;
   END_VAR
   VAR_TEMP
      TOP_SI : Struct
         EV_CLASS : Byte;
         EV_NUM : Byte;
         PRIORITY : Byte;
         NUM : Byte;
         TYP2_3 : Byte;
         TYP1 : Byte;
         ZI1 : Word;
         ZI2_3 : DWord;
      END_STRUCT;
      START_UP_SI : Struct
         EV_CLASS : Byte;
         EV_NUM : Byte;
         PRIORITY : Byte;
         NUM : Byte;
         TYP2_3 : Byte;
         TYP1 : Byte;
         ZI1 : Word;
         ZI2_3 : DWord;
      END_STRUCT;
      ERR : Int;
   END_VAR
BEGIN


   (* this FB is only necessary for siemens sps
   the siemens sps timer counts from 0 to 2^31-1 and starts at 0 sfter overrun.
   this means that the bit 31 (the highest bit ) will never be used and therefore
   a problem arises when t2 - t1 is checked.
   t2 - t1 is always valid also in an timer overrun situation where the time t1 is very high and t2 is very low.
   the result of the subtraction t2 - t1 however is still valid.
   this calculation does not work for soiemens because the highest bit is not used.

   this module stores the highest bit, changes the highest bit at every overrun occurence and stuffs ther highest bit in the output.
   the output is then used by t_plc_us and t_plc_ms.

   the correction needs and fb and not a function because the value of the highest bit has to be stored.

   do never use this function block in a codesys environment. the timer in codesys is correct and runs from 0 to 2^32-1
   *)

   (* read actual startup info *)
   (* OB1_SCAN_1  BYTE  -  B#16#01: Abschluss des Neustarts (Warmstarts)
                        -  B#16#02: Abschluss des Wiederanlaufs
                        -  B#16#03: Abschluss des freien Zyklus
                        -  B#16#04: Abschluss des Kaltstarts
                        -  B#16#05: Erster OB 1-Zyklus der neuen Master-CPU nach 
                                    Master-Reserve-Umschaltung und STOP des 
                                    bisherigen Masters *)

   #ERR := RD_SINFO (TOP_SI => #TOP_SI, START_UP_SI => #START_UP_SI);

   (* reset last_time on system startup *)
   IF #TOP_SI.EV_NUM = 1 OR #TOP_SI.EV_NUM = 2 OR #TOP_SI.EV_NUM = 4 OR NOT #init THEN 
       #last_time := 0;
       #bit31 := false;
       #init := true;
   END_IF;

   (* read the system timer *)
   #tx := DINT_TO_DWORD(T_CONV(TIME_TCK()));

   (* stuff the highest bit into the timer value *)
   #at_tx[7] := #bit31;

   (* check for overrun *)
   IF DWORD_TO_DINT(#tx) < DWORD_TO_DINT(#last_time) THEN
       (* an overrun has occured, change the value of the highest bit *)
       #bit31 := NOT #bit31;
   END_IF;

   (* stuff the highest bit into the timer value *)
   #at_tx[7] := #bit31;

   (* remember the last system time for the next overrun check *)
   #last_time := #tx;


   (* revision history
   DA  14.9.2007 rev 1.0
     original version

   DA  24.2.2008 rev 1.1
     added self reset on system startup

   DA   2.5.2008 rev 1.2
     correct a problem running under OB35

   DA  12.3.2009 rev 1.3
     correct a problem run on different CPUs

   DA  22.12.2009 rev 1.4
     correct a problem on startup

   DA  19.09.2011 rev 1.5
     correct a error in code 
   *)
END_FUNCTION_BLOCK

FUNCTION_BLOCK "TP_X"   // FB69, SCL
TITLE = TP_X
{ S7_Optimized_Access := 'FALSE' }
AUTHOR : hugo
FAMILY : GENERAT
NAME : TP_R
VERSION : 1.3
// retriggerable edge triggered pulse similar to TP but with a retrigger function
// if the pt input is 0 then output is always low.
// 
// uses: T_PLC_MS [FC64]
//       STIME [FB64],IDB_STIME [DB64]
   VAR_INPUT
      IN : Bool;
      PT : Time;
   END_VAR
   VAR_OUTPUT
      Q : Bool;
      ET : Time;
   END_VAR
   VAR
      edge : Bool;
      start : Time;
      tx : Time;
   END_VAR
   VAR_TEMP
      TOP_SI : Struct
         EV_CLASS : Byte;
         EV_NUM : Byte;
         PRIORITY : Byte;
         NUM : Byte;
         TYP2_3 : Byte;
         TYP1 : Byte;
         ZI1 : Word;
         ZI2_3 : DWord;
      END_STRUCT;
      START_UP_SI : Struct
         EV_CLASS : Byte;
         EV_NUM : Byte;
         PRIORITY : Byte;
         NUM : Byte;
         TYP2_3 : Byte;
         TYP1 : Byte;
         ZI1 : Word;
         ZI2_3 : DWord;
      END_STRUCT;
      ERR : Int;
   END_VAR
BEGIN


   (* read actual startup info *)
   (* OB1_SCAN_1  BYTE  -  B#16#01: Abschluss des Neustarts (Warmstarts)
                        -  B#16#02: Abschluss des Wiederanlaufs
                        -  B#16#03: Abschluss des freien Zyklus
                        -  B#16#04: Abschluss des Kaltstarts
                        -  B#16#05: Erster OB 1-Zyklus der neuen Master-CPU nach 
                                    Master-Reserve-Umschaltung und STOP des 
                                    bisherigen Masters *)

   #ERR := RD_SINFO (TOP_SI => #TOP_SI, START_UP_SI => #START_UP_SI);

   (* read system_time *)
   #tx := T_CONV(DWORD_TO_DINT("T_PLC_MS"()));

   (* reset last_time on system startup *)
   IF #TOP_SI.EV_NUM = 1 OR #TOP_SI.EV_NUM = 2 OR #TOP_SI.EV_NUM = 4 THEN 
       #start := #tx;
   END_IF;

   (* rising edge trigger *)
   IF #IN AND NOT #edge THEN
       #start := #tx;
       #Q := #PT > t#0ms;
   ELSIF #Q THEN
       #ET := #tx - #start;
       IF #ET >= #PT THEN
           #Q := FALSE;
           #ET := t#0ms;
       END_IF;
   END_IF;
   #edge := #IN;


   (* revision history
   hm  4. aug 2006     rev 1.0
       original version

   hm  17. sep 2007    rev 1.1
       replaced time() with T_PLC_MS() for compatibility reasons

   hm  19. oct. 2008   rev 1.2
       renamed to TP_R to TP_X for compatibility reasons

   hm  17. dec. 2008   rev 1.3
       code optimized

   *)
END_FUNCTION_BLOCK

FUNCTION_BLOCK "_RMP_B"   // FB93, SCL
TITLE = _RMP_B
{ S7_Optimized_Access := 'FALSE' }
AUTHOR : hugo
FAMILY : SIGGEN
NAME : _RMP_B
VERSION : 1.2
// _RMP_B generates a ramp on an external var of type byte
// tr is the total ramp time, E is an enable and dir the direction of the ramp
// 
// uses: T_PLC_MS [FC64]
//       STIME [FB64],IDB_STIME [DB64]
//       FRMP_B [FC424]
   VAR_INPUT
      DIR : Bool;
      "E" : Bool := TRUE;
      TR : Time;
   END_VAR
   VAR_IN_OUT
      RMP : Byte;
   END_VAR
   VAR
      tx : Time;
      tl : Time;
      tn : Time;
      init : Bool;
      last_dir : Bool;
      start : Byte;
   END_VAR
   VAR_TEMP
      TOP_SI : Struct
         EV_CLASS : Byte;
         EV_NUM : Byte;
         PRIORITY : Byte;
         NUM : Byte;
         TYP2_3 : Byte;
         TYP1 : Byte;
         ZI1 : Word;
         ZI2_3 : DWord;
      END_STRUCT;
      START_UP_SI : Struct
         EV_CLASS : Byte;
         EV_NUM : Byte;
         PRIORITY : Byte;
         NUM : Byte;
         TYP2_3 : Byte;
         TYP1 : Byte;
         ZI1 : Word;
         ZI2_3 : DWord;
      END_STRUCT;
      ERR : Int;
   END_VAR
BEGIN


   (* read actual startup info *)
   (* OB1_SCAN_1  BYTE  -  B#16#01: Abschluss des Neustarts (Warmstarts)
                        -  B#16#02: Abschluss des Wiederanlaufs
                        -  B#16#03: Abschluss des freien Zyklus
                        -  B#16#04: Abschluss des Kaltstarts
                        -  B#16#05: Erster OB 1-Zyklus der neuen Master-CPU nach 
                                    Master-Reserve-Umschaltung und STOP des 
                                    bisherigen Masters *)

   #ERR := RD_SINFO (TOP_SI => #TOP_SI, START_UP_SI => #START_UP_SI);

   (* reset last_time on system startup *)
   IF #TOP_SI.EV_NUM = 1 OR #TOP_SI.EV_NUM = 2 OR #TOP_SI.EV_NUM = 4 THEN 
       #init := false;
   END_IF;

   (* read system timer *)
   #tx := T_CONV(DWORD_TO_DINT("T_PLC_MS"()));

   IF #"E" AND #init AND (#DIR = #last_dir) AND (#RMP <> INT_TO_BYTE(DINT_TO_INT(SEL(G:=#DIR, IN0:=0, IN1:=255)))) AND #TR = #tn THEN
     #RMP := "FRMP_B"(START:=#start,DIR:=#DIR, TD:=#tx - #tl, TR:=#TR);
   ELSE
     #init := TRUE;
     #tl := #tx;
     #tn := #TR;
     #start := #RMP;
   END_IF;
   #last_dir := #DIR;



   (* revison history
   hm  22. oct. 2008 rev 1.0
     original version

   hm  20. nov. 2008 rev 1.1
     set default for E to be TRUE
     added init

   hm  19. nov. 2011 rev 1.2
     new code
   *)
END_FUNCTION_BLOCK

FUNCTION_BLOCK "_RMP_W"   // FB94, SCL
TITLE = _RMP_W
{ S7_Optimized_Access := 'FALSE' }
AUTHOR : hugo
FAMILY : SIGGEN
NAME : _RMP_W
VERSION : 1.1
// _RMP_B generates a ramp on an external var of type byte
// tr is the total ramp time, E is an enable and dir the direction of the ramp
// 
// uses: T_PLC_MS [FC64]
//       STIME [FB64],IDB_STIME [DB64]
   VAR_INPUT
      DIR : Bool;
      "E" : Bool := TRUE;
      TR : Time;
   END_VAR
   VAR_IN_OUT
      RMP : Word;
   END_VAR
   VAR
      tx : DWord;
      tl : DWord;
      "step" : DInt;
      init : Bool;
      last_dir : Bool;
   END_VAR
   VAR_TEMP
      TOP_SI : Struct
         EV_CLASS : Byte;
         EV_NUM : Byte;
         PRIORITY : Byte;
         NUM : Byte;
         TYP2_3 : Byte;
         TYP1 : Byte;
         ZI1 : Word;
         ZI2_3 : DWord;
      END_STRUCT;
      START_UP_SI : Struct
         EV_CLASS : Byte;
         EV_NUM : Byte;
         PRIORITY : Byte;
         NUM : Byte;
         TYP2_3 : Byte;
         TYP1 : Byte;
         ZI1 : Word;
         ZI2_3 : DWord;
      END_STRUCT;
      ERR : Int;
   END_VAR
BEGIN


   (* read actual startup info *)
   (* OB1_SCAN_1  BYTE  -  B#16#01: Abschluss des Neustarts (Warmstarts)
                        -  B#16#02: Abschluss des Wiederanlaufs
                        -  B#16#03: Abschluss des freien Zyklus
                        -  B#16#04: Abschluss des Kaltstarts
                        -  B#16#05: Erster OB 1-Zyklus der neuen Master-CPU nach 
                                    Master-Reserve-Umschaltung und STOP des 
                                    bisherigen Masters *)

   #ERR := RD_SINFO (TOP_SI => #TOP_SI, START_UP_SI => #START_UP_SI);

   (* reset last_time on system startup *)
   IF #TOP_SI.EV_NUM = 1 OR #TOP_SI.EV_NUM = 2 OR #TOP_SI.EV_NUM = 4 THEN 
       #init := FALSE;
   END_IF;

   #tx := "T_PLC_MS"();
   IF #"E" AND #init THEN
       (* we need to set tl = tx when direction changes *)
       IF #DIR XOR #last_dir THEN
        #tl := #tx;
        #last_dir := #DIR;
       END_IF;
       (* check_elapsed time and calculate only if necessary *)
       IF #TR > t#0s THEN
           #"step" := DWORD_TO_DINT(SHL(IN:=DINT_TO_DWORD(DWORD_TO_DINT(#tx)-DWORD_TO_DINT(#tl)), N:=16)) / T_CONV(#TR);
       ELSE
           #"step" := 65535;
       END_IF;
       IF #"step" > 0 THEN
           (* perform the step on the ramp *)
           #tl := #tx;
           (* calculate the step response *)
           IF NOT #DIR THEN #"step" := - #"step"; END_IF;
           #RMP := DINT_TO_WORD(LIMIT(MN:=0, IN:=WORD_TO_DINT(#RMP) + #"step", MX:=65535));
       END_IF;
   ELSE
       #tl := #tx;
       #init := TRUE;
   END_IF;


   (* revison history
   hm  22. oct. 2008   rev 1.0
       original version

   hm  20. nov. 2008   rev 1.1
       set default for E to be TRUE
       added init

   *)
END_FUNCTION_BLOCK

FUNCTION_BLOCK "GEN_PULSE"   // FB95, SCL
TITLE = GEN_PULSE
{ S7_Optimized_Access := 'FALSE' }
AUTHOR : hugo
FAMILY : SIGGEN
NAME : GEN_PULS
VERSION : 1.5
// GEN_PULSE uses the internal sps time to generate a continuous output waveform with programmable high and low time.
// clk_prg depending on the accuracy of the system clock.
// when time is 0 the high and low times are exactly one cycle.
// ENQ = TRUE will start and ENQ = FALSE will stop the generator.
// 
// uses: T_PLC_MS [FC64]
//       STIME [FB64],IDB_STIME [DB64]
   VAR_INPUT
      ENQ : Bool := TRUE;
      PTH : Time;
      PTL : Time;
   END_VAR
   VAR_OUTPUT
      Q : Bool;
   END_VAR
   VAR
      tx : Time;
      tn : Time;
      init : Bool;
   END_VAR
   VAR_TEMP
      TOP_SI : Struct
         EV_CLASS : Byte;
         EV_NUM : Byte;
         PRIORITY : Byte;
         NUM : Byte;
         TYP2_3 : Byte;
         TYP1 : Byte;
         ZI1 : Word;
         ZI2_3 : DWord;
      END_STRUCT;
      START_UP_SI : Struct
         EV_CLASS : Byte;
         EV_NUM : Byte;
         PRIORITY : Byte;
         NUM : Byte;
         TYP2_3 : Byte;
         TYP1 : Byte;
         ZI1 : Word;
         ZI2_3 : DWord;
      END_STRUCT;
      ERR : Int;
   END_VAR
BEGIN


     (* read actual startup info *)
     (* OB1_SCAN_1  BYTE  -  B#16#01: Abschluss des Neustarts (Warmstarts)
                          -  B#16#02: Abschluss des Wiederanlaufs
                          -  B#16#03: Abschluss des freien Zyklus
                          -  B#16#04: Abschluss des Kaltstarts
                          -  B#16#05: Erster OB 1-Zyklus der neuen Master-CPU nach 
                                      Master-Reserve-Umschaltung und STOP des 
                                      bisherigen Masters *)

     #ERR := RD_SINFO (TOP_SI => #TOP_SI, START_UP_SI => #START_UP_SI);

     (* reset last_time on system startup *)
     IF #TOP_SI.EV_NUM = 1 OR #TOP_SI.EV_NUM = 2 OR #TOP_SI.EV_NUM = 4 THEN 
       #init := FALSE;
     END_IF;

     IF #ENQ THEN
       #tx := T_CONV(DWORD_TO_DINT("T_PLC_MS"()));
       IF NOT #init THEN #init := TRUE; #tn := #tx; END_IF;
       IF #tx - #tn >= SEL(G:=#Q, IN0:=#PTL, IN1:=#PTH) THEN
         #tn := #tn + SEL(G:=#Q, IN0:=#PTL, IN1:=#PTH);
         #Q := NOT #Q;
       END_IF;
     ELSE
       #Q := FALSE;
       #init := FALSE;
     END_IF;


   (* revision history
   hm  29. jun. 2008 rev 1.0
     original version

   hm 23. nov. 2008 rev 1.1
     set default for enq to be true

   hm  18. jul. 2009 rev 1.2
     improved performance

   hm  13. nov. 2009 rev 1.3
     corrected error

   hm  16. feb. 2011 rev 1.4
     corrected an error when timer overflows

   hm  8. apr. 2011  rev 1.5
     ptl and pth was exchanged
   *)
END_FUNCTION_BLOCK

FUNCTION_BLOCK "GEN_PW2"   // FB96, SCL
TITLE = GEN_PW2
{ S7_Optimized_Access := 'FALSE' }
AUTHOR : hugo
FAMILY : SIGGEN
NAME : GEN_PW2